screen "Statie Hidraulica" 1920x1080, template "Template_1"
   Rectangle "Rectangle_26" at 1435,281 size 25x72
      Appearance <- "DB_Inspect_Pistoane_Piston_1"
   SymbolLibrary "Symbol library_12" at 919,817 size 79x75
      on Click: SetTag("DB_Inspect_Pistoane_PompaC", 0)
      Appearance <- "DB_Status_Pistoane_Status_Piston_C"
   SymbolLibrary "Symbol library_13" at 992,840 size 110x71
      Appearance <- "DB_Status_Pistoane_Status_Piston_C"
   GraphicView "Graphic view_21" at 894,866 size 56x21; Picture "Graphic_102"
      Appearance <- "DB_Inspect_Pistoane_Piston_1"
   SymbolLibrary "Symbol library_5" at 925,709 size 79x75
      Appearance <- "DB_Status_Pistoane_Status_Piston_C"
      on Click: SetTag("DB_Inspect_Pistoane_PompaC", 0)
   SymbolLibrary "Symbol library_4" at 925,601 size 79x75
      Appearance <- "DB_Status_Pistoane_Status_Piston_B"
      on Click: SetTag("DB_Inspect_Pistoane_PompaB", 0)
   SymbolLibrary "Symbol library_3" at 925,493 size 79x75
      Appearance <- "DB_Status_Pistoane_Status_Piston_A"
      on Click: SetTag("DB_Inspect_Pistoane_PompaA", 0)
   SymbolLibrary "Symbol library_8" at 927,385 size 77x74
      Appearance <- "DB_Status_Pistoane_Status_Pison_2"
      on Click: SetTag("DB_Inspect_Pistoane_Pompa2", 0)
   SymbolLibrary "Symbol library_1" at 923,279 size 79x75
      Appearance <- "DB_Inspect_Pistoane_Pompa1"
      on Press: SetTag("DB_Inspect_Pistoane_Pompa1", 0)
   Bar "Bar_6" at 1163,534 size 102x44; MinimumValue 0
      ProcessValue <- "DB_Inspect_Pistoane_Presiune_1"
   TextField "Text field_3" at 26,401 size 265x38; Text 'Oil Volume / Ölvolumen'
   TextField "Text field_2" at 20,878 size 364x38; Text 'Oil Temperature / Öltemperatur'
   Switch "Switch_2" at 560,308 size 173x84; TextOn 'Piston 1 / Kolben 1'; CaptionText 'Switch'; TextOff 'Piston 1 / Kolben 1'
      on SwitchOn: SetTag("DB_Inspect_Pistoane_Piston_2", 0); SetTag("DB_Inspect_Pistoane_Piston_A", 0); SetTag("DB_Inspect_Pistoane_Piston_B", 0); SetTag("DB_Inspect_Pistoane_Piston_C", 0)
      Appearance <- "DB_Inspect_Pistoane_Piston_1"
      ProcessValue <- "DB_Inspect_Pistoane_Piston_1"
   Switch "Switch_3" at 562,410 size 173x84; TextOn 'Piston 2 / Kolben 2'; CaptionText 'Switch'; TextOff 'Piston 2 / Kolben 2'
      on SwitchOn: SetTag("DB_Inspect_Pistoane_Piston_1", 0); SetTag("DB_Inspect_Pistoane_Piston_A", 0); SetTag("DB_Inspect_Pistoane_Piston_B", 0); SetTag("DB_Inspect_Pistoane_Piston_C", 0)
      Appearance <- "DB_Inspect_Pistoane_Piston_2"
      ProcessValue <- "DB_Inspect_Pistoane_Piston_2"
   Switch "Switch_4" at 560,502 size 173x84; TextOn 'Piston A / Kolben A'; CaptionText 'Switch'; TextOff 'Piston A / Kolben A'
      on SwitchOn: SetTag("DB_Inspect_Pistoane_Piston_1", 0); SetTag("DB_Inspect_Pistoane_Piston_2", 0); SetTag("DB_Inspect_Pistoane_Piston_B", 0); SetTag("DB_Inspect_Pistoane_Piston_C", 0)
      Appearance <- "DB_Inspect_Pistoane_Piston_A"
      ProcessValue <- "DB_Inspect_Pistoane_Piston_A"
   Switch "Switch_5" at 560,604 size 173x84; TextOn 'Piston B / Kolben B'; CaptionText 'Switch'; TextOff 'Piston B / Kolben B'
      on SwitchOn: SetTag("DB_Inspect_Pistoane_Piston_2", 0); SetTag("DB_Inspect_Pistoane_Piston_A", 0); SetTag("DB_Inspect_Pistoane_Piston_1", 0); SetTag("DB_Inspect_Pistoane_Piston_C", 0)
      Appearance <- "DB_Inspect_Pistoane_Piston_B"
      ProcessValue <- "DB_Inspect_Pistoane_Piston_B"
   Switch "Switch_6" at 560,702 size 173x84; TextOn 'Piston C / Kolben C'; CaptionText 'Switch'; TextOff 'Piston C / Kolben C'
      on SwitchOn: SetTag("DB_Inspect_Pistoane_Piston_2", 0); SetTag("DB_Inspect_Pistoane_Piston_A", 0); SetTag("DB_Inspect_Pistoane_Piston_B", 0); SetTag("DB_Inspect_Pistoane_Piston_1", 0)
      Appearance <- "DB_Inspect_Pistoane_Piston_C"
      ProcessValue <- "DB_Inspect_Pistoane_Piston_C"
   Rectangle "Rectangle_8" at 754,320 size 82x63
      Appearance <- "DB_Status_Pistoane_Status_Piston_1"
   Rectangle "Rectangle_30" at 758,418 size 82x63
      Appearance <- "DB_Status_Pistoane_Status_Pison_2"
   Rectangle "Rectangle_9" at 756,512 size 82x63
      Appearance <- "DB_Status_Pistoane_Status_Piston_A"
   Rectangle "Rectangle_10" at 756,610 size 82x63
      Appearance <- "DB_Status_Pistoane_Status_Piston_B"
   Rectangle "Rectangle_37" at 756,710 size 82x63
      Appearance <- "DB_Status_Pistoane_Status_Piston_C"
   Switch "Switch_7" at 596,204 size 226x98; CaptionText 'Switch'; TextOff 'Piston Status Kolben Status'; TextOn 'Piston Status Kolben Status'
   Button "Button_3" at 262,707 size 192x68; TextOff 'Set T=0C / Stellen Sie T=0C'
      on Release: SetTag("DB_HMI_Set_T0", 0)
      on Press: SetTag("DB_HMI_Set_T0", 1)
   Button "Button_4" at 262,628 size 192x68; TextOff 'Set T=50C / Stellen Sie T=50C'
      on Release: SetTag("DB_HMI_Set_T50", 0)
      on Press: SetTag("DB_HMI_Set_T50", 1)
   Bar "Bar_1" at 28,514 size 116x350; MinimumValue 0; MaximumValue 50
      ProcessValue <- "DB_HMI_Temp_Ulei"
   Rectangle "Rectangle_2" at 178,333 size 106x50
      Appearance <- "DB_HMI_Volum_Ulei"
   Bar "Bar_3" at 38,56 size 106x345; MinimumValue 0; MaximumValue 50
      ProcessValue <- "DB_HMI_Volum_Ulei"
   Button "Button_1" at 190,140 size 63x64; TextOff '+'
      on Release: SetTag("DB_HMI_Add_Ulei", 0)
      on Press: SetTag("DB_HMI_Add_Ulei", 1)
      Appearance <- "DB_HMI_Volum_Ulei"
   Rectangle "Rectangle_1" at 170,56 size 113x50
      Appearance <- "DB_HMI_Volum_Ulei"
   TextField "Text field_1" at 184,332 size 121x38; Text 'MIN'
      Appearance <- "DB_HMI_Volum_Ulei"
   Button "Button_2" at 190,262 size 63x64; TextOff 'Text'
      on Release: SetTag("DB_HMI_Sub_Ulei", 0)
      on Press: SetTag("DB_HMI_Sub_Ulei", 1)
      Appearance <- "DB_HMI_Volum_Ulei"
   TextField "Text field_13" at 178,56 size 125x38; Text 'MAX'
      Appearance <- "DB_HMI_Volum_Ulei"
   GraphicView "Graphic view_24" at 1305,408 size 146x23; Picture "Graphic_102"
      Appearance <- "DB_Inspect_Pistoane_Piston_1"
   GraphicView "Graphic view_28" at 1105,392 size 221x84; Picture "Graphic_65"
      Appearance <- "DB_Inspect_Pistoane_Piston_1"
   GraphicView "Graphic view_29" at 1305,516 size 146x23; Picture "Graphic_102"
      Appearance <- "DB_Inspect_Pistoane_Piston_1"
   GraphicView "Graphic view_33" at 1105,500 size 221x84; Picture "Graphic_65"
      Appearance <- "DB_Inspect_Pistoane_Piston_1"
   GraphicView "Graphic view_34" at 1305,624 size 146x23; Picture "Graphic_102"
      Appearance <- "DB_Inspect_Pistoane_Piston_1"
   GraphicView "Graphic view_35" at 900,650 size 56x21; Picture "Graphic_102"
      Appearance <- "DB_Inspect_Pistoane_Piston_1"
   GraphicView "Graphic view_38" at 1105,608 size 221x84; Picture "Graphic_65"
      Appearance <- "DB_Inspect_Pistoane_Piston_1"
   GraphicView "Graphic view_39" at 1305,732 size 146x23; Picture "Graphic_102"
      Appearance <- "DB_Inspect_Pistoane_Piston_1"
   GraphicView "Graphic view_40" at 900,758 size 56x21; Picture "Graphic_102"
      Appearance <- "DB_Inspect_Pistoane_Piston_1"
   GraphicView "Graphic view_43" at 1105,716 size 221x84; Picture "Graphic_65"
      Appearance <- "DB_Inspect_Pistoane_Piston_1"
   TextField "Text field_5" at 1177,297 size 95x22; Text 'Presiune / Druck'
   TextField "Text field_4" at 1176,401 size 92x22; Text 'Pressure / Druck'
   TextField "Text field_6" at 1177,511 size 100x22; Text 'Pressure / Druck'
   TextField "Text field_7" at 1177,617 size 100x22; Text 'Pressure / Druck'
   TextField "Text field_8" at 1177,725 size 100x22; Text 'Pressure / Druck'
   IOField "I/O field_1" at 1165,328 size 96x32; FormatPattern 9999999
   GraphicView "Graphic view_19" at 1303,302 size 146x23; Picture "Graphic_102"
      Appearance <- "DB_Inspect_Pistoane_Piston_1"
   GraphicView "Graphic view_23" at 1103,286 size 221x84; Picture "Graphic_65"
      Appearance <- "DB_Inspect_Pistoane_Piston_1"
   TextField "Text field_10" at 1176,294 size 92x22; Text 'Pressure / Druck'
   Bar "Bar_4" at 1163,424 size 102x44; MinimumValue 0
      ProcessValue <- "DB_Inspect_Pistoane_Presiune_2"
   Bar "Bar_5" at 1166,532 size 102x44; MinimumValue 0
      ProcessValue <- "DB_Inspect_Pistoane_Presiune_A"
   Bar "Bar_7" at 1163,641 size 102x44; MinimumValue 0
      ProcessValue <- "DB_Inspect_Pistoane_Presiune_B"
   Bar "Bar_8" at 1163,748 size 102x44; MinimumValue 0
      ProcessValue <- "DB_Inspect_Pistoane_Presiune_C"
   Bar "Bar_10" at 1163,318 size 102x44; MinimumValue 0
      ProcessValue <- "DB_Inspect_Pistoane_Presiune_1"
   GraphicView "Graphic view_49" at 880,252 size 35x653; Picture "Graphic_110"
   GraphicView "Graphic view_11" at 358,466 size 135x135; Picture "Graphic_97"
      Visibility <- "DB_HMI_Status_Incalzire/Racire_Ulei"
   GraphicView "Graphic view_7" at 363,472 size 122x126; Picture "Graphic_93"
      Visibility <- "DB_HMI_Ventilator_Cald"
   GraphicView "Graphic view_6" at 367,472 size 117x126; Picture "Graphic_92"
      Visibility <- "DB_HMI_Ventilator_Cald"
   GraphicView "Graphic view_8" at 364,476 size 120x118; Picture "Graphic_94"
      Visibility <- "DB_HMI_Ventilator_Cald"
   GraphicView "Graphic view_9" at 360,473 size 124x122; Picture "Graphic_95"
      Visibility <- "DB_HMI_Ventilator_Cald"
   GraphicView "Graphic view_13" at 358,466 size 135x136; Picture "Graphic_98"
      Visibility <- "DB_HMI_Status_Incalzire/Racire_Ulei"
   GraphicView "Graphic view_14" at 367,476 size 120x118; Picture "Graphic_96"
      Visibility <- "DB_HMI_Status_Incalzire/Racire_Ulei"
   GraphicView "Graphic view_16" at 358,467 size 134x134; Picture "Graphic_98"
      Visibility <- "DB_HMI_Status_Incalzire/Racire_Ulei"
   GraphicView "Graphic view_10" at 222,468 size 134x134; Picture "Graphic_61"
      Visibility <- "DB_HMI_Status_Incalzire/Racire_Ulei"
   GraphicView "Graphic view_1" at 232,474 size 116x120; Picture "Graphic_49"
      Visibility <- "DB_HMI_Ventilator_Rece"
   GraphicView "Graphic view_2" at 228,474 size 121x125; Picture "Graphic_50"
      Visibility <- "DB_HMI_Ventilator_Rece"
   GraphicView "Graphic view_3" at 228,477 size 121x118; Picture "Graphic_51"
      Visibility <- "DB_HMI_Ventilator_Rece"
   GraphicView "Graphic view_5" at 226,475 size 122x121; Picture "Graphic_52"
      Visibility <- "DB_HMI_Ventilator_Rece"
   GraphicView "Graphic view_4" at 222,468 size 134x134; Picture "Graphic_98"
      Visibility <- "DB_HMI_Status_Incalzire/Racire_Ulei"
   GraphicView "Graphic view_12" at 230,478 size 120x118; Picture "Graphic_96"
      Visibility <- "DB_HMI_Status_Incalzire/Racire_Ulei"
   GraphicView "Graphic view_17" at 223,467 size 134x134; Picture "Graphic_98"
      Visibility <- "DB_HMI_Status_Incalzire/Racire_Ulei"
   GraphicView "Graphic view_18" at 230,476 size 120x118; Picture "Graphic_96"
      Visibility <- "DB_HMI_Status_Incalzire/Racire_Ulei"
   SymbolLibrary "Symbol library_7" at 885,192 size 66x76
      Appearance <- "DB_Inspect_Pistoane_PompaPrincipala"
   GraphicView "Graphic view_30" at 900,542 size 55x21; Picture "Graphic_102"
      Appearance <- "DB_Inspect_Pistoane_Piston_1"
   GraphicView "Graphic view_25" at 900,434 size 56x21; Picture "Graphic_102"
      Appearance <- "DB_Inspect_Pistoane_Piston_1"
   GraphicView "Graphic view_20" at 901,328 size 53x21; Picture "Graphic_102"
      Appearance <- "DB_Inspect_Pistoane_Piston_1"
   GraphicView "Graphic view_15" at 366,474 size 120x118; Picture "Graphic_96"
      Visibility <- "DB_HMI_Status_Incalzire/Racire_Ulei"
   SymbolLibrary "Symbol library_2" at 995,302 size 110x71
      Appearance <- "DB_Status_Pistoane_Status_Piston_1"
   SymbolLibrary "Symbol library_6" at 998,407 size 110x71
      Appearance <- "DB_Status_Pistoane_Status_Pison_2"
   SymbolLibrary "Symbol library_9" at 998,516 size 110x71
      Appearance <- "DB_Status_Pistoane_Status_Piston_A"
   SymbolLibrary "Symbol library_10" at 998,624 size 110x71
      Appearance <- "DB_Status_Pistoane_Status_Piston_B"
   SymbolLibrary "Symbol library_11" at 998,732 size 110x71
      Appearance <- "DB_Status_Pistoane_Status_Piston_C"
   Button "Button_7" at 1344,200 size 118x40; TextOff 'Fix'
      on Activate: SetTag("DB_Inspect_Pistoane_Pompa1", 2); SetTag("DB_Inspect_Pistoane_Pompa2", 2); SetTag("DB_Inspect_Pistoane_PompaA", 2); SetTag("DB_Inspect_Pistoane_PompaB", 2); SetTag("DB_Inspect_Pistoane_PompaC", 2); SetTag("DB_Inspect_Pistoane_StatusPump1", 1)
   Button "Button_8" at 1344,143 size 118x40; TextOff 'Jinx P1'
      on Activate: SetTag("DB_Inspect_Pistoane_Pompa1", 0); SetTag("DB_Inspect_Pistoane_StatusPump1", 0)
   Switch "Switch_9" at 562,808 size 173x84; TextOn 'Piston 3 / Kolben C'; CaptionText 'Switch'; TextOff 'Piston 3 / Kolben C'
      on SwitchOn: SetTag("DB_Inspect_Pistoane_Piston_2", 0); SetTag("DB_Inspect_Pistoane_Piston_A", 0); SetTag("DB_Inspect_Pistoane_Piston_B", 0); SetTag("DB_Inspect_Pistoane_Piston_1", 0)
   GraphicView "Graphic view_22" at 1299,842 size 146x23; Picture "Graphic_102"
      Appearance <- "DB_Inspect_Pistoane_Piston_1"
   GraphicView "Graphic view_26" at 1099,826 size 221x84; Picture "Graphic_65"
      Appearance <- "DB_Inspect_Pistoane_Piston_1"
   Bar "Bar_2" at 1157,858 size 102x44; MinimumValue 0
      ProcessValue <- "DB_Inspect_Pistoane_Presiune_C"
   Rectangle "Rectangle_7" at 1437,387 size 25x72
      Appearance <- "DB_Inspect_Pistoane_Piston_2"
   Rectangle "Rectangle_19" at 1437,495 size 25x72
      Appearance <- "DB_Inspect_Pistoane_Piston_A"
   Rectangle "Rectangle_25" at 1437,603 size 25x72
      Appearance <- "DB_Inspect_Pistoane_Piston_B"
   Rectangle "Rectangle_36" at 1437,711 size 25x72
      Appearance <- "DB_Inspect_Pistoane_Piston_C"
   Rectangle "Rectangle_44" at 1433,817 size 25x72
      Appearance <- "DB_Inspect_Pistoane_Piston_C"
   Group "Group" at 1435,281 size 58x158

screen "Log_Cutii" 1920x1080, template "Template_1"
   on GenerateScreen: "VBFunction_2"()
   Rectangle "Rectangle_9" at 16,165 size 1422x79
      Appearance <- "Viz_Pachet_1"
   Rectangle "Rectangle_10" at 16,307 size 1422x77
      Appearance <- "Viz_Pachet_3"
   Rectangle "Rectangle_13" at 16,727 size 1422x77
      Appearance <- "Viz_Pachet_9"
   Rectangle "Rectangle_12" at 16,586 size 1422x81
      Appearance <- "Viz_Pachet_7"
   Rectangle "Rectangle_11" at 16,445 size 1422x80
      Appearance <- "Viz_Pachet_5"
   Rectangle "Rectangle_7" at 16,803 size 1422x65
      Appearance <- "Viz_Pachet_10"
   Rectangle "Rectangle_6" at 16,665 size 1422x64
      Appearance <- "Viz_Pachet_8"
   Rectangle "Rectangle_5" at 16,524 size 1422x64
      Appearance <- "Viz_Pachet_6"
   Rectangle "Rectangle_4" at 16,383 size 1422x64
      Appearance <- "Viz_Pachet_4"
   Rectangle "Rectangle_3" at 16,243 size 1422x65
      Appearance <- "Viz_Pachet_2"
   TextField "Text field_4" at 256,122 size 57x34; Text 'ID'
   TextField "Text field_2" at 830,122 size 152x34; Text 'Weight / Gewicht'
   TextField "Text field_3" at 1236,122 size 227x34; Text 'Destination / Ziel'
   TextField "Text field_5" at 1008,122 size 243x34; Text 'Gearbox type'
   Button "Button_6" at 28,530 size 132x52; TextOff 'Details / Einzelheiten'
      on Click: InvertBit("Viz_Pachet_6"); "VBFunction_1"(5); "VBFunction_5"(); SetTag("Viz_Pachet_2", 0); SetTag("Viz_Pachet_3", 0); SetTag("Viz_Pachet_4", 0); SetTag("Viz_Pachet_5", 0); SetTag("Viz_Pachet_1", 0); SetTag("Viz_Pachet_7", 0); SetTag("Viz_Pachet_8", 0); SetTag("Viz_Pachet_9", 0); SetTag("Viz_Pachet_10", 0); function_efd93a16("Pop-up screen_1", 0, 0, 0, -1, 1)
   IOField "I/O field_5" at 186,178 size 173x52; FormatPattern 999
      ProcessValue <- "[0]"
      Appearance <- "Viz_Pachet_1"
   IOField "I/O field_6" at 366,176 size 477x52; FormatPattern 9999999999999999999999999999999999999999
      ProcessValue <- "[0]"
      Appearance <- "Viz_Pachet_1"
   Button "Button_3" at 26,178 size 132x52; TextOff 'Details / Einzelheiten'
      on Click: InvertBit("Viz_Pachet_1"); "VBFunction_1"(0); "VBFunction_5"(); SetTag("Viz_Pachet_2", 0); SetTag("Viz_Pachet_3", 0); SetTag("Viz_Pachet_4", 0); SetTag("Viz_Pachet_5", 0); SetTag("Viz_Pachet_6", 0); SetTag("Viz_Pachet_7", 0); SetTag("Viz_Pachet_8", 0); SetTag("Viz_Pachet_9", 0); SetTag("Viz_Pachet_10", 0); function_efd93a16("Pop-up screen_1", 0, 0, 0, -1, 1)
   IOField "I/O field_7" at 819,179 size 173x52; FormatPattern 999
      Visibility <- "Viz_Pachet_1"
      ProcessValue <- "Greutate_TEST"
      Appearance <- "Viz_Pachet_1"
   IOField "I/O field_8" at 1048,178 size 173x52; FormatPattern ????????????????????????????????????????????????????????????????????????????????
      Visibility <- "Viz_Pachet_1"
      ProcessValue <- "Tip_TEST"
      Appearance <- "Viz_Pachet_1"
   IOField "I/O field_9" at 1244,178 size 173x52; FormatPattern ????????????????????????????????????????????????????????????????????????????????
      Visibility <- "Viz_Pachet_1"
      ProcessValue <- "Destinatie_TEST"
      Appearance <- "Viz_Pachet_1"
   IOField "I/O field_20" at 191,249 size 173x52; FormatPattern 999
      ProcessValue <- "[1]"
      Appearance <- "Viz_Pachet_2"
   IOField "I/O field_21" at 373,247 size 477x52; FormatPattern 9999999999999999999999999999999999999999
      ProcessValue <- "[1]"
      Appearance <- "Viz_Pachet_2"
   Button "Button_14" at 28,250 size 132x52; TextOff 'Details / Einzelheiten'
      on Click: InvertBit("Viz_Pachet_2"); "VBFunction_1"(1); "VBFunction_5"(); SetTag("Viz_Pachet_1", 0); SetTag("Viz_Pachet_3", 0); SetTag("Viz_Pachet_4", 0); SetTag("Viz_Pachet_5", 0); SetTag("Viz_Pachet_6", 0); SetTag("Viz_Pachet_7", 0); SetTag("Viz_Pachet_8", 0); SetTag("Viz_Pachet_9", 0); SetTag("Viz_Pachet_10", 0); function_efd93a16("Pop-up screen_1", 0, 0, 0, -1, 1)
   IOField "I/O field_22" at 818,249 size 173x52; FormatPattern 999
      Visibility <- "Viz_Pachet_2"
      ProcessValue <- "Greutate_TEST"
      Appearance <- "Viz_Pachet_2"
   IOField "I/O field_23" at 1049,249 size 173x52; FormatPattern ????????????????????????????????????????????????????????????????????????????????
      Visibility <- "Viz_Pachet_2"
      ProcessValue <- "Tip_TEST"
      Appearance <- "Viz_Pachet_2"
   IOField "I/O field_24" at 1244,250 size 173x52; FormatPattern ????????????????????????????????????????????????????????????????????????????????
      Visibility <- "Viz_Pachet_2"
      ProcessValue <- "Destinatie_TEST"
      Appearance <- "Viz_Pachet_2"
   IOField "I/O field_25" at 190,319 size 173x52; FormatPattern 999
      ProcessValue <- "[2]"
      Appearance <- "Viz_Pachet_3"
   IOField "I/O field_26" at 370,317 size 477x52; FormatPattern 9999999999999999999999999999999999999999
      ProcessValue <- "[2]"
      Appearance <- "Viz_Pachet_3"
   Button "Button_15" at 26,316 size 132x52; TextOff 'Details / Einzelheiten'
      on Click: InvertBit("Viz_Pachet_3"); "VBFunction_1"(2); "VBFunction_5"(); SetTag("Viz_Pachet_2", 0); SetTag("Viz_Pachet_1", 0); SetTag("Viz_Pachet_4", 0); SetTag("Viz_Pachet_5", 0); SetTag("Viz_Pachet_6", 0); SetTag("Viz_Pachet_7", 0); SetTag("Viz_Pachet_8", 0); SetTag("Viz_Pachet_9", 0); SetTag("Viz_Pachet_10", 0); function_efd93a16("Pop-up screen_1", 0, 0, 0, -1, 1)
   IOField "I/O field_27" at 818,814 size 173x52; FormatPattern 999
      Visibility <- "Viz_Pachet_10"
      ProcessValue <- "Greutate_TEST"
      Appearance <- "Viz_Pachet_10"
   IOField "I/O field_28" at 1043,806 size 173x52; FormatPattern ????????????????????????????????????????????????????????????????????????????????
      Visibility <- "Viz_Pachet_10"
      ProcessValue <- "Tip_TEST"
      Appearance <- "Viz_Pachet_10"
   IOField "I/O field_29" at 1239,806 size 173x52; FormatPattern ????????????????????????????????????????????????????????????????????????????????
      Visibility <- "Viz_Pachet_10"
      ProcessValue <- "Destinatie_TEST"
      Appearance <- "Viz_Pachet_10"
   IOField "I/O field_10" at 186,390 size 173x52; FormatPattern 999
      ProcessValue <- "[3]"
      Appearance <- "Viz_Pachet_4"
   IOField "I/O field_11" at 371,389 size 477x52; FormatPattern 9999999999999999999999999999999999999999
      ProcessValue <- "[3]"
      Appearance <- "Viz_Pachet_4"
   Button "Button_4" at 28,390 size 132x52; TextOff 'Details / Einzelheiten'
      on Click: InvertBit("Viz_Pachet_4"); "VBFunction_1"(3); "VBFunction_5"(); SetTag("Viz_Pachet_2", 0); SetTag("Viz_Pachet_3", 0); SetTag("Viz_Pachet_1", 0); SetTag("Viz_Pachet_5", 0); SetTag("Viz_Pachet_6", 0); SetTag("Viz_Pachet_7", 0); SetTag("Viz_Pachet_8", 0); SetTag("Viz_Pachet_9", 0); SetTag("Viz_Pachet_10", 0); function_efd93a16("Pop-up screen_1", 0, 0, 0, -1, 1)
   IOField "I/O field_12" at 819,323 size 173x52; FormatPattern 999
      ProcessValue <- "Greutate_TEST"
      Visibility <- "Viz_Pachet_3"
      Appearance <- "Viz_Pachet_3"
   IOField "I/O field_13" at 1044,315 size 173x52; FormatPattern ????????????????????????????????????????????????????????????????????????????????
      ProcessValue <- "Tip_TEST"
      Visibility <- "Viz_Pachet_3"
      Appearance <- "Viz_Pachet_3"
   IOField "I/O field_14" at 1245,315 size 173x52; FormatPattern ????????????????????????????????????????????????????????????????????????????????
      ProcessValue <- "Destinatie_TEST"
      Visibility <- "Viz_Pachet_3"
      Appearance <- "Viz_Pachet_3"
   IOField "I/O field_15" at 186,460 size 173x52; FormatPattern 999
      ProcessValue <- "[4]"
      Appearance <- "Viz_Pachet_5"
   IOField "I/O field_16" at 366,458 size 477x52; FormatPattern 9999999999999999999999999999999999999999
      ProcessValue <- "[4]"
      Appearance <- "Viz_Pachet_5"
   Button "Button_5" at 28,460 size 132x52; TextOff 'Details / Einzelheiten'
      on Click: InvertBit("Viz_Pachet_5"); "VBFunction_1"(4); "VBFunction_5"(); SetTag("Viz_Pachet_2", 0); SetTag("Viz_Pachet_3", 0); SetTag("Viz_Pachet_4", 0); SetTag("Viz_Pachet_1", 0); SetTag("Viz_Pachet_6", 0); SetTag("Viz_Pachet_7", 0); SetTag("Viz_Pachet_8", 0); SetTag("Viz_Pachet_9", 0); SetTag("Viz_Pachet_10", 0); function_efd93a16("Pop-up screen_1", 0, 0, 0, -1, 1)
   IOField "I/O field_17" at 819,393 size 173x52; FormatPattern 999
      Visibility <- "Viz_Pachet_4"
      ProcessValue <- "Greutate_TEST"
      Appearance <- "Viz_Pachet_4"
   IOField "I/O field_18" at 1044,385 size 173x52; FormatPattern ????????????????????????????????????????????????????????????????????????????????
      Visibility <- "Viz_Pachet_4"
      ProcessValue <- "Tip_TEST"
      Appearance <- "Viz_Pachet_4"
   IOField "I/O field_19" at 1240,385 size 173x52; FormatPattern ????????????????????????????????????????????????????????????????????????????????
      Visibility <- "Viz_Pachet_4"
      ProcessValue <- "Destinatie_TEST"
      Appearance <- "Viz_Pachet_4"
   IOField "I/O field_30" at 186,530 size 173x52; FormatPattern 999
      ProcessValue <- "[5]"
      Appearance <- "Viz_Pachet_6"
   IOField "I/O field_31" at 366,528 size 477x52; FormatPattern 9999999999999999999999999999999999999999
      ProcessValue <- "[5]"
      Appearance <- "Viz_Pachet_6"
   IOField "I/O field_32" at 818,460 size 173x52; FormatPattern 999
      Visibility <- "Viz_Pachet_5"
      ProcessValue <- "Greutate_TEST"
      Appearance <- "Viz_Pachet_5"
   IOField "I/O field_35" at 1046,454 size 173x52; FormatPattern ????????????????????????????????????????????????????????????????????????????????
      Visibility <- "Viz_Pachet_5"
      ProcessValue <- "Tip_TEST"
      Appearance <- "Viz_Pachet_5"
   IOField "I/O field_36" at 1240,455 size 173x52; FormatPattern ????????????????????????????????????????????????????????????????????????????????
      Visibility <- "Viz_Pachet_5"
      ProcessValue <- "Destinatie_TEST"
      Appearance <- "Viz_Pachet_5"
   IOField "I/O field_37" at 186,600 size 173x52; FormatPattern 999
      ProcessValue <- "[6]"
      Appearance <- "Viz_Pachet_7"
   IOField "I/O field_38" at 366,598 size 477x52; FormatPattern 9999999999999999999999999999999999999999
      ProcessValue <- "[6]"
      Appearance <- "Viz_Pachet_7"
   Button "Button_7" at 28,600 size 132x52; TextOff 'Details / Einzelheiten'
      on Click: InvertBit("Viz_Pachet_7"); "VBFunction_1"(6); "VBFunction_5"(); SetTag("Viz_Pachet_2", 0); SetTag("Viz_Pachet_3", 0); SetTag("Viz_Pachet_4", 0); SetTag("Viz_Pachet_5", 0); SetTag("Viz_Pachet_6", 0); SetTag("Viz_Pachet_1", 0); SetTag("Viz_Pachet_8", 0); SetTag("Viz_Pachet_9", 0); SetTag("Viz_Pachet_10", 0); function_efd93a16("Pop-up screen_1", 0, 0, 0, -1, 1)
   IOField "I/O field_39" at 819,533 size 173x52; FormatPattern 999
      Visibility <- "Viz_Pachet_6"
      ProcessValue <- "Greutate_TEST"
      Appearance <- "Viz_Pachet_6"
   IOField "I/O field_40" at 1044,525 size 173x52; FormatPattern ????????????????????????????????????????????????????????????????????????????????
      Visibility <- "Viz_Pachet_6"
      ProcessValue <- "Tip_TEST"
      Appearance <- "Viz_Pachet_6"
   IOField "I/O field_41" at 1247,525 size 173x52; FormatPattern ????????????????????????????????????????????????????????????????????????????????
      Visibility <- "Viz_Pachet_6"
      ProcessValue <- "Destinatie_TEST"
      Appearance <- "Viz_Pachet_6"
   IOField "I/O field_42" at 186,670 size 173x52; FormatPattern 999
      ProcessValue <- "[7]"
      Appearance <- "Viz_Pachet_8"
   IOField "I/O field_43" at 366,668 size 477x52; FormatPattern 9999999999999999999999999999999999999999
      ProcessValue <- "[7]"
      Appearance <- "Viz_Pachet_8"
   Button "Button_8" at 28,670 size 132x52; TextOff 'Details / Einzelheiten'
      on Click: InvertBit("Viz_Pachet_8"); "VBFunction_1"(7); "VBFunction_5"(); SetTag("Viz_Pachet_2", 0); SetTag("Viz_Pachet_3", 0); SetTag("Viz_Pachet_1", 0); SetTag("Viz_Pachet_5", 0); SetTag("Viz_Pachet_6", 0); SetTag("Viz_Pachet_7", 0); SetTag("Viz_Pachet_1", 0); SetTag("Viz_Pachet_9", 0); SetTag("Viz_Pachet_10", 0); function_efd93a16("Pop-up screen_1", 0, 0, 0, -1, 1)
   IOField "I/O field_44" at 819,603 size 173x52; FormatPattern 999
      Visibility <- "Viz_Pachet_7"
      ProcessValue <- "Greutate_TEST"
      Appearance <- "Viz_Pachet_7"
   IOField "I/O field_45" at 1044,595 size 173x52; FormatPattern ????????????????????????????????????????????????????????????????????????????????
      Visibility <- "Viz_Pachet_7"
      ProcessValue <- "Tip_TEST"
      Appearance <- "Viz_Pachet_7"
   IOField "I/O field_46" at 1240,595 size 173x52; FormatPattern ????????????????????????????????????????????????????????????????????????????????
      Visibility <- "Viz_Pachet_7"
      ProcessValue <- "Destinatie_TEST"
      Appearance <- "Viz_Pachet_7"
   IOField "I/O field_47" at 186,740 size 173x52; FormatPattern 999
      ProcessValue <- "[8]"
      Appearance <- "Viz_Pachet_9"
   IOField "I/O field_48" at 366,738 size 477x52; FormatPattern 9999999999999999999999999999999999999999
      ProcessValue <- "[8]"
      Appearance <- "Viz_Pachet_9"
   Button "Button_16" at 28,740 size 132x52; TextOff 'Details / Einzelheiten'
      on Click: InvertBit("Viz_Pachet_9"); "VBFunction_1"(8); "VBFunction_5"(); SetTag("Viz_Pachet_2", 0); SetTag("Viz_Pachet_3", 0); SetTag("Viz_Pachet_4", 0); SetTag("Viz_Pachet_5", 0); SetTag("Viz_Pachet_6", 0); SetTag("Viz_Pachet_7", 0); SetTag("Viz_Pachet_8", 0); SetTag("Viz_Pachet_1", 0); SetTag("Viz_Pachet_10", 0); function_efd93a16("Pop-up screen_1", 0, 0, 0, -1, 1)
   IOField "I/O field_49" at 819,673 size 173x52; FormatPattern 999
      Visibility <- "Viz_Pachet_8"
      ProcessValue <- "Greutate_TEST"
      Appearance <- "Viz_Pachet_8"
   IOField "I/O field_50" at 1039,673 size 173x52; FormatPattern ????????????????????????????????????????????????????????????????????????????????
      Visibility <- "Viz_Pachet_8"
      ProcessValue <- "Tip_TEST"
      Appearance <- "Viz_Pachet_8"
   IOField "I/O field_51" at 1242,670 size 173x52; FormatPattern ????????????????????????????????????????????????????????????????????????????????
      Visibility <- "Viz_Pachet_8"
      ProcessValue <- "Destinatie_TEST"
      Appearance <- "Viz_Pachet_8"
   IOField "I/O field_52" at 186,810 size 173x52; FormatPattern 999
      ProcessValue <- "[9]"
      Appearance <- "Viz_Pachet_10"
   IOField "I/O field_53" at 366,808 size 477x52; FormatPattern 9999999999999999999999999999999999999999
      ProcessValue <- "[9]"
      Appearance <- "Viz_Pachet_10"
   Button "Button_17" at 28,810 size 132x52; TextOff 'Details / Einzelheiten'
      on Click: InvertBit("Viz_Pachet_10"); "VBFunction_1"(9); "VBFunction_5"(); SetTag("Viz_Pachet_2", 0); SetTag("Viz_Pachet_3", 0); SetTag("Viz_Pachet_4", 0); SetTag("Viz_Pachet_5", 0); SetTag("Viz_Pachet_6", 0); SetTag("Viz_Pachet_7", 0); SetTag("Viz_Pachet_8", 0); SetTag("Viz_Pachet_9", 0); SetTag("Viz_Pachet_1", 0); function_efd93a16("Pop-up screen_1", 0, 0, 0, -1, 1)
   IOField "I/O field_54" at 819,743 size 173x52; FormatPattern 999
      Visibility <- "Viz_Pachet_9"
      ProcessValue <- "Greutate_TEST"
      Appearance <- "Viz_Pachet_9"
   IOField "I/O field_55" at 1042,740 size 173x52; FormatPattern ????????????????????????????????????????????????????????????????????????????????
      Visibility <- "Viz_Pachet_9"
      ProcessValue <- "Tip_TEST"
      Appearance <- "Viz_Pachet_9"
   IOField "I/O field_56" at 1240,735 size 173x52; FormatPattern ????????????????????????????????????????????????????????????????????????????????
      Visibility <- "Viz_Pachet_9"
      ProcessValue <- "Destinatie_TEST"
      Appearance <- "Viz_Pachet_9"
   TextField "Text field_6" at 539,120 size 106x34; Text 'Data / Datum'
   Button "Button_1" at 1639,335 size 250x88; TextOff 'Show QR / QR anzeigen'
      on Click: function_efd93a16("Pop-up screen_1", 1640, 450, -1, 2, 0)
      ObjectEnable <- "QR_En"

PopupScreen "Pop-up screen_1" 250x250
   HTMLBrowser "HTML browser_1" at 8,13 size 225x225

screen "AdminPage" 1920x1080, template "Template_1"
   Button "Button_1" at 126,88 size 258x76; TextOff 'Shift details / Schichtdetails'
      on Click: SetTag("DB_HMI_Detalii_Cutii", 1); SetTag("DB_HMI_Modificare_Param", 0); SetTag("DB_HMI_Sistem_Racire", 0)
      Appearance <- "DB_HMI_Detalii_Cutii"
   Button "Button_3" at 52,188 size 401x76; TextOff 'Packets parameters / Paketparameter'
      on Click: SetTag("DB_HMI_Detalii_Cutii", 0); SetTag("DB_HMI_Sistem_Racire", 0); SetTag("DB_HMI_Modificare_Param", 1)
      Appearance <- "DB_HMI_Modificare_Param"
   DateTimeField "Date/time field_1" at 636,1 size 888x47
   Rectangle "Rectangle_2" at 502,58 size 1150x244
      Visibility <- "DB_HMI_Detalii_Cutii"
   TextField "Text field_16" at 453,79 size 1193x52; Text 'Packets in the last 24 hours / Pakete in den letzten 24 Stunden'
      Visibility <- "DB_HMI_Detalii_Cutii"
   TextField "Text field_17" at 513,150 size 373x52; Text 'Total Packets / Gesamtpakete'
      Visibility <- "DB_HMI_Detalii_Cutii"
   TextField "Text field_18" at 877,149 size 305x52; Text 'Shift 1 / Schicht 1'
      Visibility <- "DB_HMI_Detalii_Cutii"
   TextField "Text field_19" at 1134,150 size 305x52; Text 'Shift 2 / Schicht 2'
      Visibility <- "DB_HMI_Detalii_Cutii"
   TextField "Text field_20" at 1381,150 size 305x52; Text 'Shift 3 / Schicht 3'
      Visibility <- "DB_HMI_Detalii_Cutii"
   IOField "I/O field_10" at 561,211 size 186x82; FormatPattern 999
      Visibility <- "DB_HMI_Detalii_Cutii"
      ProcessValue <- "DB_HMI_Total_Packets"
   IOField "I/O field_11" at 905,216 size 186x82; FormatPattern 999
      Visibility <- "DB_HMI_Detalii_Cutii"
      ProcessValue <- "DB_HMI_Pachete_Schimb1"
   IOField "I/O field_12" at 1157,216 size 186x82; FormatPattern 999
      Visibility <- "DB_HMI_Detalii_Cutii"
      ProcessValue <- "DB_HMI_Pachete_Schimb2"
   Rectangle "Rectangle_6" at 501,312 size 1150x589
      Visibility <- "DB_HMI_Detalii_Cutii"
   TrendView "Trend view_1" at 524,331 size 1123x563
      Visibility <- "DB_HMI_Detalii_Cutii"
   IOField "I/O field_13" at 1406,216 size 186x82; FormatPattern 999
      Visibility <- "DB_HMI_Detalii_Cutii"
      ProcessValue <- "DB_HMI_Pachete_Schimb3"
   Button "Button_2" at 52,297 size 401x76; TextOff 'Cooling parameters / Kühlparameter'
      on Click: SetTag("DB_HMI_Detalii_Cutii", 0); SetTag("DB_HMI_Sistem_Racire", 1); SetTag("DB_HMI_Modificare_Param", 0)
      Appearance <- "DB_HMI_Sistem_Racire"
   Button "Button_4" at 138,824 size 219x76; TextOff 'Log Out / Ausloggen'
      on Click: ActivateScreen("Home", 0)
   Rectangle "Rectangle_5" at 502,313 size 1150x511
      Visibility <- "DB_HMI_Modificare_Param"
   Rectangle "Rectangle_3" at 502,58 size 1150x244
      Visibility <- "DB_HMI_Modificare_Param"
   IOField "I/O field_1" at 524,199 size 186x82; Authorization "Monitor"; FormatPattern 999; Unit  kg
      ProcessValue <- "DB_general_GreutateManual"
      Visibility <- "DB_HMI_Modificare_Param"
   TextField "Text field_1" at 632,88 size 816x100; Text 'Nominal weights for gearboxes / Nenngewichte für Getriebe'
      Visibility <- "DB_HMI_Modificare_Param"
   TextField "Text field_2" at 432,151 size 370x40; Text 'Manual / Schalt'
      Visibility <- "DB_HMI_Modificare_Param"
   IOField "I/O field_2" at 781,203 size 186x82; FormatPattern 999; Unit  kg
      ProcessValue <- "DB_general_GreutateAutomata"
      Visibility <- "DB_HMI_Modificare_Param"
   TextField "Text field_3" at 674,150 size 370x40; Text 'Automatic / Automatik'
      Visibility <- "DB_HMI_Modificare_Param"
   TextField "Text field_4" at 1031,131 size 713x112; Text 'Weight tolerance percentage / Prozentsatz der Gewichtstoleranz'
      Visibility <- "DB_HMI_Modificare_Param"
   IOField "I/O field_3" at 1228,203 size 186x82; FormatPattern 99; Unit  %
      Visibility <- "DB_HMI_Modificare_Param"
      ProcessValue <- "DB_general_Procent_Toleranta"
   TextField "Text field_6" at 687,327 size 593x52; Text 'Truck parameters / LKW-Parameter'
      Visibility <- "DB_HMI_Modificare_Param"
   TextField "Text field_7" at 512,386 size 253x52; Text 'Truck A / LKW A'
      Visibility <- "DB_HMI_Modificare_Param"
   TextField "Text field_8" at 910,386 size 301x52; Text 'Truck B / LKW B'
      Visibility <- "DB_HMI_Modificare_Param"
   TextField "Text field_9" at 1371,386 size 253x52; Text 'Truck C / LKW C'
      Visibility <- "DB_HMI_Modificare_Param"
   TextField "Text field_10" at 494,453 size 341x76; Text 'Max Load / Tragfähigkeit'
      Visibility <- "DB_HMI_Modificare_Param"
   IOField "I/O field_4" at 560,523 size 186x82; Authorization "Monitor"; FormatPattern 999; Unit  kg
      Visibility <- "DB_HMI_Modificare_Param"
      ProcessValue <- "DB_HMI_MaxLoad_A"
   IOField "I/O field_7" at 972,521 size 186x82; Authorization "Monitor"; FormatPattern 999; Unit  kg
      Visibility <- "DB_HMI_Modificare_Param"
      ProcessValue <- "DB_HMI_MaxLoad_B"
   IOField "I/O field_8" at 1406,522 size 186x82; Authorization "Monitor"; FormatPattern 999; Unit  kg
      Visibility <- "DB_HMI_Modificare_Param"
      ProcessValue <- "DB_HMI_MaxLoad_C"
   TextField "Text field_13" at 504,608 size 385x76; Text 'Expected quantity / Erwartete Menge'
      Visibility <- "DB_HMI_Modificare_Param"
   IOField "I/O field_5" at 560,675 size 186x82; Authorization "Monitor"; FormatPattern 99
      Visibility <- "DB_HMI_Modificare_Param"
      ProcessValue <- "Locuri_A"
   IOField "I/O field_6" at 975,671 size 186x82; Authorization "Monitor"; FormatPattern 99
      Visibility <- "DB_HMI_Modificare_Param"
      ProcessValue <- "Locuri_B"
   IOField "I/O field_9" at 1406,672 size 186x82; Authorization "Monitor"; FormatPattern 99
      Visibility <- "DB_HMI_Modificare_Param"
      ProcessValue <- "Locuri_C"
   TextField "Text field_14" at 888,608 size 385x76; Text 'Expected quantity / Erwartete Menge'
      Visibility <- "DB_HMI_Modificare_Param"
   TextField "Text field_15" at 1295,608 size 385x76; Text 'Expected quantity / Erwartete Menge'
      Visibility <- "DB_HMI_Modificare_Param"
   TextField "Text field_11" at 919,449 size 341x76; Text 'Max Load / Tragfähigkeit'
      Visibility <- "DB_HMI_Modificare_Param"
   TextField "Text field_12" at 1357,447 size 332x76; Text 'Max Load / Tragfähigkeit'
      Visibility <- "DB_HMI_Modificare_Param"
   Rectangle "Rectangle_7" at 501,58 size 1150x244
      Visibility <- "DB_HMI_Sistem_Racire"
   Rectangle "Rectangle_8" at 501,312 size 1150x589
      Visibility <- "DB_HMI_Sistem_Racire"
   TrendView "Trend view_2" at 511,331 size 1123x563
      Visibility <- "DB_HMI_Sistem_Racire"
   TextField "Text field_5" at 503,77 size 1105x52; Text 'Parameters of the cooling sysytem / Parameter des Kühlsystems'
      Visibility <- "DB_HMI_Sistem_Racire"
   TextField "Text field_21" at 694,131 size 601x52; Text 'Temp Max'
      Visibility <- "DB_HMI_Sistem_Racire"
   TextField "Text field_22" at 326,131 size 591x52; Text 'Temp Min'
      Visibility <- "DB_HMI_Sistem_Racire"
   TextField "Text field_24" at 1046,134 size 640x52; Text 'Temp Optim'
      Visibility <- "DB_HMI_Sistem_Racire"
   IOField "I/O field_14" at 557,199 size 186x82; Authorization "Monitor"; FormatPattern 99; Unit  C
      ProcessValue <- "DB_HMI_Temp_Min"
      Visibility <- "DB_HMI_Sistem_Racire"
   IOField "I/O field_15" at 942,200 size 186x82; Authorization "Monitor"; FormatPattern 99; Unit  C
      ProcessValue <- "DB_HMI_Temp_Max"
      Visibility <- "DB_HMI_Sistem_Racire"
   IOField "I/O field_16" at 1306,202 size 186x82; Authorization "Monitor"; FormatPattern 99; Unit  C
      ProcessValue <- "DB_HMI_Temp_Optim"
      Visibility <- "DB_HMI_Sistem_Racire"

screen "ServerTeste" 1920x1080
   TextField "Text field_1" at 343,298 size 144x22; Text 'Inmatriculare TIR:'

PopupScreen "Pop-up screen_2" 240x240
   TextField "Text field_1" at 65,89 size 15x22; Text 'Text'
   TextField "Text field_2" at 23,37 size 120x22; Text 'Total weight / Gesamtgewicht'
   TextField "Text field_3" at 23,79 size 140x22; Text 'Available places / Verfügbare Plätze'
   IOField "I/O field_1" at 169,35 size 50x32; FormatPattern 999
   IOField "I/O field_2" at 169,79 size 50x32; FormatPattern 999

VB script "VBFunction_2"
   'Select din SQL
   Dim con,rs
   Dim DataTimp
   Dim value
   Dim paddingSpace
   Dim rezultate
   Dim ids,greutate, destinatie, tipCutie
   Set con=CreateObject("adodb.connection")
   Set rs=CreateObject("adodb.recordset")
   
   Dim i
   i=0
   
   con.open"Driver={MySQL ODBC 8.0 Unicode Driver};Server=localhost:3306;Database=colete;User=root;Password=;Option=3;"
   rs.open "select * from pachete ORDER BY ID DESC Limit 10",con
   rs.MoveFirst
   
   While Not rs.EOF
       SmartTags("Array_Id")(i) = rs.Fields(0) 
       SmartTags("Array_Data")(i) = rs.Fields(4) 
       rs.MoveNext
       i = i +1
   Wend
   
   
   	
   con.Close

VB script "VBFunction_4"
   'Insert in SQL
   
   
   
   If SmartTags("RdyToLog") = True Then
   Dim con,rs
   Dim value
   Dim paddingSpace
   Dim rezultate
   
   
   
   
   Dim greutate, destinatie, tipCutie
   Set greutate = SmartTags("DB_HMI_Greutate")
   Set destinatie = SmartTags("Destinatie_Pachet")
   Set tipCutie = SmartTags("Tip_Cutie_Pachet")
   ' cod nou-----------------------
   
   
   'Dim Timp
   'Timp = Time
   'Dim TimpStamp
   Dim dtsnow
   Dim dd, mm, yy, hh, nn, ss
   Dim DataValue, TimpValue
   Dim dtsvalue
   dtsnow = Now()
   dd = Right("00" & Day(dtsnow), 2)
   mm = Right("00" & Month(dtsnow), 2)
   yy = Year(dtsnow)
   hh = Right("00" & Hour(dtsnow), 2)
   nn = Right("00" & Minute(dtsnow), 2)
   ss = Right("00" & Second(dtsnow), 2)
   
   'Build the date string in the format yyyy-mm-dd
   DataValue = yy & "-" & mm & "-" & dd
   'Build the time string in the format hh:mm:ss
   TimpValue = hh & ":" & nn & ":" & ss
   'Concatenate both together to build the timestamp yyyy-mm-dd hh:mm:ss
   dtsvalue = DataValue & " " & TimpValue
   
   'Dim Data
   'Data = Date
   
   
   'Dim Timp
   'Timp = Time
   'Dim TimpStamp
   
   Dim stringlog, delimitator
   
   'delimitator = " "
   'TimpStamp= Data & delimitator & Timp
   
   delimitator = " - "
   
   stringlog =greutate & delimitator & destinatie & delimitator & tipCutie & delimitator & dtsvalue
   
   
   Set con=CreateObject("adodb.connection")
   Set rs=CreateObject("adodb.recordset")
   Dim sqlString, partSql
   partSql= "INSERT INTO colete.pachete (Greutate,Destinatie,Tip,Data) VALUES ('"
   
   sqlString=partSql & greutate 
   
   partSql="','"
   sqlString=sqlString & partSql & destinatie & partSql & tipCutie  & partSql & dtsvalue
   
   partSql="')"
   
   sqlString=sqlString & partSql
   
   con.open"Driver={MySQL ODBC 8.0 Unicode Driver};Server=localhost:3306;Database=colete;User=root;Password=;Option=3;"
   rs.open sqlString,con
   
   con.Close
   
   
   Set sqlString = Nothing
   
   
   'resetam rdy to log ul
   
   Dim val 
   val = False
   SmartTags("RdyToLog") = val
   
   
   
   
   End If

VB script "VBFunction_6"
   'Tip:
   ' 1. Use the <CTRL+SPACE> or <CTRL+I> shortcut to open a list of all objects and functions
   ' 2. Write the code using the HMI Runtime object.
   '  Example: HmiRuntime.Screens("Screen_1").
   ' 3. Use the <CTRL+J> shortcut to create an object reference.
   'Write the code as of this position:
   
   'Dim runphp
   'Set runphp = CreateObject("wscript.shell")
   'runphp.Run"C:\xampp\htdocs\Test_Qr\cronjob.bat",7
   
   
   
   Dim url
    url = "http://localhost/Test_Qr/test.php?id=2"
   SmartTags("url") = url

VB script "VBFunction_5"
   'Tip:
   ' 1. Use the <CTRL+SPACE> or <CTRL+I> shortcut to open a list of all objects and functions
   ' 2. Write the code using the HMI Runtime object.
   '  Example: HmiRuntime.Screens("Screen_1").
   ' 3. Use the <CTRL+J> shortcut to create an object reference.
   'Write the code as of this position:
   
   
   'REFRESH
   
   Dim fileobj,file,path, rezultate
   Set fileobj=CreateObject("Scripting.FileSystemObject")
   ' How to write file
   path="C:\xampp\htdocs\Test_QR_V02\Test\Test\DATEQR.txt"
   
   Dim tip, destinatie
   
   'Select Case SmartTags("Destinatie_Pachet")
   '	Case 1
   '		destinatie = "Locatie A"
   '	Case 2
   '		destinatie = "Locatie B"
   '	Case 3
   '		destinatie = "Locatie C"
   '	Case Else
   '		destinatie = "Destinatie necunoscuta"
   'End Select
   '
   'Select Case SmartTags("Tip_Cutie_Pachet")
   '	Case 1
   '		tip = "Automata"
   '	Case 2
   '		tip = "Manuala"
   '	Case Else
   '		tip = "Destinatie necunoscuta"
   'End Select
   '''
   rezultate = "Id Colet: " & SmartTags("ID_TEST") & vbCrLf  & "Greutate Colet: " & SmartTags("Greutate_TEST") & vbCrLf & "Destinatie Colet: " & SmartTags("Destinatie_TEST") & vbCrLf & "Tip Colet: " & SmartTags("Tip_TEST") & vbCrLf & "Data Colet: " & SmartTags("Data") 
    
   Set file = fileobj.CreateTextFile(path,True)
   file.Write rezultate
   file.Close
   
   Set fileobj = Nothing
   
   Dim updateqr
   Set updateqr = CreateObject("wscript.shell")
   updateqr.Run "C:\xampp\htdocs\Test_QR_V02\Test\Test\callqr.bat",7
   
   SmartTags("QR_En") = True

VB script "VBFunction_1"
   'Tip:
   ' 1. Use the <CTRL+SPACE> or <CTRL+I> shortcut to open a list of all objects and functions
   ' 2. Write the code using the HMI Runtime object.
   '  Example: HmiRuntime.Screens("Screen_1").
   ' 3. Use the <CTRL+J> shortcut to create an object reference.
   'Write the code as of this position:
   
   
   'Select din SQL
   
   
   Dim con,rs
   Dim destinatie, tipCutie
   Set con=CreateObject("adodb.connection")
   Set rs=CreateObject("adodb.recordset")
   
   
   
   
   Dim fileobj,file,path, rezultate
   Set fileobj=CreateObject("Scripting.FileSystemObject")
   ' How to write file
   path="C:\xampp\htdocs\Test_QR_V02\Test\Test\DATEQR.txt"
   
   
   con.open"Driver={MySQL ODBC 8.0 Unicode Driver};Server=localhost:3306;Database=colete;User=root;Password=;Option=3;"
   rs.open "select * from pachete WHERE ID = " & SmartTags("Array_Id")(id) & " ORDER BY ID DESC Limit 1",con
   'rs.MoveFirst
   
   'While Not rs.EOF
      
   tipCutie = rs.Fields(3) 
   destinatie = rs.Fields(2) 
   SmartTags("Greutate_TEST") = rs.Fields(1) 
   SmartTags("ID_TEST") = rs.Fields(0) 
   SmartTags("Data") = rs.Fields(4) 
   'Wend
   
   
   
   
   Select Case destinatie
   	Case 1
   		SmartTags("Destinatie_TEST") = "Location A"
   	Case 2
   		SmartTags("Destinatie_TEST") = "Location B"
   	Case 3
   		SmartTags("Destinatie_TEST") = "Location C"
   	Case Else
   		SmartTags("Destinatie_TEST") = "Destination unknown"
   End Select
   
   Select Case tipCutie
   	Case 2
   		SmartTags("Tip_TEST") = "Automatic"
   	Case 1
   		SmartTags("Tip_TEST") = "Manual"
   	Case Else
   		SmartTags("Tip_TEST") = "Destination unknown"
   End Select
   
   rezultate = "Id Colet: " & SmartTags("ID_TEST") & vbCrLf  & "Greutate Colet: " & SmartTags("Greutate_TEST") & vbCrLf & "Destinatie Colet: " & SmartTags("Destinatie_TEST") & vbCrLf & "Tip Colet: " & SmartTags("Tip_TEST") & vbCrLf & "Data Colet: " & SmartTags("Data") 
    
   Set file = fileobj.CreateTextFile(path,True)
   file.Write rezultate
   file.Close
   
   Set fileobj = Nothing
   
   Dim updateqr
   Set updateqr = CreateObject("wscript.shell")
   updateqr.Run "C:\xampp\htdocs\Test_QR_V02\Test\Test\callqr.bat",7
   
   con.Close
*)